   
   			//Position x (Forward)
    			IF NOT IN_xLastModalityLoadBkw AND NOT IN_xLastModalityUnloadBkw THEN
   				//Tail
   				IF TMP_dCap = 0 THEN
   					Scada_Plate[IN_iIndexArray, TMP_dCap, TMP_dLite].dTail_PosX_mm := TMP_dHeadPosition_mm - (IN_tPlate.rgtCap[TMP_dCap].dLength_cmm / 100);
   				ELSE
   					Scada_Plate[IN_iIndexArray, TMP_dCap, TMP_dLite].dTail_PosX_mm := Scada_Plate[IN_iIndexArray, TMP_dCap - 1, TMP_dLite].dTail_PosX_mm -
   					(IN_tPlate.rgtCap[TMP_dCap].dLength_cmm / 100) - (IN_tPlate.rgtCap[TMP_dCap-1].dReqGapForConv_cmm /100);	//(IN_tPlate.dGapCaps_cmm / 100);
   				END_IF;
   				//Head
   				Scada_Plate[IN_iIndexArray, TMP_dCap, TMP_dLite].dHead_PosX_mm := TMP_dHeadPosition_mm;
   				IF TMP_dCap > 0 THEN
   					Scada_Plate[IN_iIndexArray, TMP_dCap, TMP_dLite].dHead_PosX_mm := Scada_Plate[IN_iIndexArray, TMP_dCap - 1, TMP_dLite].dHead_PosX_mm -
   					(IN_tPlate.rgtCap[TMP_dCap - 1].dLength_cmm / 100) - (IN_tPlate.rgtCap[TMP_dCap-1].dReqGapForConv_cmm /100);	//(IN_tPlate.dGapCaps_cmm / 100);
   				END_IF;
   			END_IF;
   			//Position x (Backward)
   			//Head
   			IF IN_xLastModalityLoadBkw OR IN_xLastModalityUnloadBkw THEN
   				//  Head
   				IF TMP_dCap = 0 THEN
   					Scada_Plate[IN_iIndexArray, TMP_dCap, TMP_dLite].dHead_PosX_mm := TMP_dConveyorLenght - TMP_dHeadPosition_mm + (IN_tPlate.dLength_cmm / 100);
   				ELSE
   					Scada_Plate[IN_iIndexArray, TMP_dCap, TMP_dLite].dHead_PosX_mm := (TMP_dConveyorLenght - TMP_dHeadPosition_mm
   					+ (IN_tPlate.dLength_cmm / 100)) - (IN_tPlate.rgtCap[TMP_dCap - 1].dLength_cmm / 100) - (IN_tPlate.rgtCap[TMP_dCap-1].dReqGapForConv_cmm /100);	//(IN_tPlate.dGapCaps_cmm / 100);
   				END_IF;
   				//  Tail
   				IF TMP_dCap = 0 THEN
   					Scada_Plate[IN_iIndexArray, TMP_dCap, TMP_dLite].dTail_PosX_mm :=
   					Scada_Plate[IN_iIndexArray, TMP_dCap, TMP_dLite].dHead_PosX_mm - (IN_tPlate.rgtCap[TMP_dCap].dLength_cmm / 100);
   				ELSE
   					Scada_Plate[IN_iIndexArray, TMP_dCap, TMP_dLite].dTail_PosX_mm :=
   					Scada_Plate[IN_iIndexArray, TMP_dCap, TMP_dLite].dHead_PosX_mm - (IN_tPlate.rgtCap[TMP_dCap].dLength_cmm / 100);
   				END_IF;
   			END_IF;
   			//Position Y
   			//Baricentre not used, without inversion (IN Fc)
   			IF NOT IN_xYWithBaricentre AND NOT IN_xYInversionLite THEN
   				IF TMP_dLite < 1 THEN
   					Scada_Plate[IN_iIndexArray, TMP_dCap, TMP_dLite].dPositionY_mm :=
   					((TMP_dWidth_mm / 2) - (IN_tPlate.rgtCap[TMP_dCap].dWidth_cmm / 100) / 2);
   				END_IF;
   			END_IF;
   			//Baricentre not used, with inversion (IN Fc)
   			IF NOT IN_xYWithBaricentre AND IN_xYInversionLite THEN
   				IF TMP_dLite < 1 THEN
   					Scada_Plate[IN_iIndexArray, TMP_dCap, TMP_dLite].dPositionY_mm :=
   					(TMP_dWidth_mm / 2) + ((IN_tPlate.rgtCap[TMP_dCap].dWidth_cmm / 100) / 2) -
   					(IN_tPlate.rgtCap[TMP_dCap].rgtLite[TMP_dLite].dWidth_cmm / 100);
   				ELSE
   					Scada_Plate[IN_iIndexArray, TMP_dCap, TMP_dLite].dPositionY_mm := Scada_Plate[IN_iIndexArray, TMP_dCap, TMP_dLite - 1].dPositionY_mm
   					- (IN_tPlate.rgtCap[TMP_dCap].rgtLite[TMP_dLite].dWidth_cmm / 100) -
   					(IN_tPlate.rgtCap[TMP_dCap-1].dReqGapForConv_cmm /100);	//(IN_tPlate.rgtCap[TMP_dCap].dGap_cmm / 100);
   				END_IF;
   			END_IF;
   			//Baricentre used, without inversion (IN Fc)
   			IF IN_xYWithBaricentre AND NOT IN_xYInversionLite THEN
   				Scada_Plate[IN_iIndexArray, TMP_dCap, TMP_dLite].dPositionY_mm :=
   				(TMP_dWidth_mm / 2) - ((IN_tPlate.rgtCap[TMP_dCap].rgtLite[TMP_dLite].dWidth_cmm / 100) / 2)
   				+ (IN_tPlate.rgtCap[TMP_dCap].rgtLite[TMP_dLite].dBarycenter_cmm / 100);
   			END_IF;
   			//Baricentre used, with inversion (IN Fc)
   			IF IN_xYWithBaricentre AND IN_xYInversionLite THEN    //Baricentre used,  inversion
   				Scada_Plate[IN_iIndexArray, TMP_dCap, TMP_dLite].dPositionY_mm :=
   				(TMP_dWidth_mm / 2) - ((IN_tPlate.rgtCap[TMP_dCap].rgtLite[TMP_dLite].dWidth_cmm / 100) / 2)
   				- (IN_tPlate.rgtCap[TMP_dCap].rgtLite[TMP_dLite].dBarycenter_cmm / 100);
   			END_IF;
   		END_IF;
   	END_FOR;
   END_FOR;
   
END_ROUTINE
END_ADD_ON_INSTRUCTION

ADD_ON_INSTRUCTION GP_SpaceConvUtilities_V1   (* revision 1.0 *)
VAR_IN_OUT
   Conveyor : SpaceConv_Utilities; {required}
   Previus_Conveyor : SpaceConv_Utilities; {required}
   Next_Conveyor : SpaceConv_Utilities; {required}
END_VAR
VAR_INPUT
   In_dModality : DINT; {required}   // Call modality 1=GlsPos|2=PrstH|3=PrstT|4=SyncH_T|5=StartLoadForward|6=StartUnloadForward|7=PrstLoad/Unload12=PrstHInversionRun|13=PrstTInversionRun |15=StartLoadBackward|16=StartUnloadBackward
END_VAR
VAR
   TMP_dVirtualSyncroPos_cmm : DINT; {access None}
   TMP_rSP_Speed_mm_min : REAL; {access None}
   TMP_rScan_ms : REAL; {access None}
   TMP_xRunning : BOOL; {access None}
   TMP_rStepAcc_mm_min : REAL; {access None}
   TMP_rLimAcc_mm_min : REAL; {access None}
   TMP_rStepDec_mm_min : REAL; {access None}
   TMP_rLimDec_mm_min : REAL; {access None}
   TMP_dRampSpace_cmm : DINT; {access None}
   TMP_dAcc_ms2 : DINT; {access None}
   TMP_dSincrhoPhotocelPos : DINT; {access None}
   TMP_dRealSpeed : REAL; {access None}
END_VAR

ROUTINE Logic   (* structured text *)
   
   CASE In_dModality OF
       2: //Preset head position
           Conveyor.O_rHeadPosition_cmm := Conveyor.CONF_MD2_MD3_dPrstPos_cmm;
           Conveyor.O_dHeadPosition_cmm := Conveyor.CONF_MD2_MD3_dPrstPos_cmm;
   
       3: //Preset Tail position
           Conveyor.O_rTailPosition_cmm := Conveyor.CONF_MD2_MD3_dPrstPos_cmm;
           Conveyor.O_dTailPosition_cmm := Conveyor.CONF_MD2_MD3_dPrstPos_cmm;
   
       4://Glass syncrhonization
           // Calculate Ramp Space
           TMP_dAcc_ms2 := Conveyor.CONST_rAcceleration_ms2 * 1000.0;
           TMP_dRampSpace_cmm := ((Conveyor.ST_dRealSpeed_mm_min / 60) * (Conveyor.ST_dRealSpeed_mm_min / 60)) / (2 * TMP_dAcc_ms2) * 100;
           TMP_dSincrhoPhotocelPos := TMP_dRampSpace_cmm + Conveyor.CONST_dSyncroPhPosition_cmm;
           CASE Conveyor.CONST_dSyncMode OF
               0://No syncro
                   Conveyor.O_xPlateSynchronized := 1;
   
               1://Syncro on head
                   IF Conveyor.ST_OS_xSynchroPhotocellHead AND NOT (Conveyor.O_xPlateSynchronized)
                       AND Conveyor.O_dHeadPosition_cmm >= TMP_dSincrhoPhotocelPos - (Conveyor.CONST_dSyncroPhWindow_cmm / 2)
                       AND Conveyor.O_dHeadPosition_cmm <= TMP_dSincrhoPhotocelPos + (Conveyor.CONST_dSyncroPhWindow_cmm / 2) THEN
                       Conveyor.O_dHeadPosition_cmm := TMP_dSincrhoPhotocelPos;
                       Conveyor.O_rHeadPosition_cmm := Conveyor.O_dHeadPosition_cmm;
                       Conveyor.O_xPlateSynchronized := 1;
                   END_IF;
               2://Syncro on tail
                   TMP_dVirtualSyncroPos_cmm := TMP_dSincrhoPhotocelPos + Conveyor.CONF_MD4_MD6_dLength_cmm;
                   IF Conveyor.ST_OS_xSynchroPhotocellTail AND NOT (Conveyor.O_xPlateSynchronized)
                       AND Conveyor.O_dHeadPosition_cmm >= TMP_dVirtualSyncroPos_cmm - (Conveyor.CONST_dSyncroPhWindow_cmm / 2)
                       AND Conveyor.O_dHeadPosition_cmm <= TMP_dVirtualSyncroPos_cmm + (Conveyor.CONST_dSyncroPhWindow_cmm / 2) THEN
                       Conveyor.O_dHeadPosition_cmm := TMP_dVirtualSyncroPos_cmm;
                       Conveyor.O_rHeadPosition_cmm := Conveyor.O_dHeadPosition_cmm;
                       Conveyor.O_xPlateSynchronized := 1;
                   END_IF;
           END_CASE;
       5://Start load
           Conveyor.O_dHeadPosition_cmm := Previus_Conveyor.O_dHeadPosition_cmm - Previus_Conveyor.CONST_dConveyorLength_cmm;
           Conveyor.O_rHeadPosition_cmm := Conveyor.O_dHeadPosition_cmm;
           Conveyor.ST_rSpeedIncrementH_mm_min := Previus_Conveyor.ST_rSpeedIncrementH_mm_min;
           Conveyor.ST_xLastModLoadBkw := 0;
           Conveyor.ST_xLastModUnloadBkw := 0;
       6://Start unload
           Conveyor.O_dTailPosition_cmm := Conveyor.O_dHeadPosition_cmm - Conveyor.CONF_MD4_MD6_dLength_cmm;
           Conveyor.O_rTailPosition_cmm := Conveyor.O_dTailPosition_cmm;
           Conveyor.ST_xLastModLoadBkw := 0;
           Conveyor.ST_xLastModUnloadBkw := 0;
       7://Load and unload simultaneous
           TMP_dAcc_ms2 := Conveyor.CONST_rAcceleration_ms2 * 1000.0;
           TMP_dRampSpace_cmm := ((Conveyor.ST_dRealSpeed_mm_min / 60) * (Conveyor.ST_dRealSpeed_mm_min / 60)) / (2 * TMP_dAcc_ms2) * 100;
           Conveyor.O_dPresetLoadUnload_cmm := ((Conveyor.CONST_dConveyorLength_cmm + TMP_dRampSpace_cmm - Conveyor.ST_dStopLoadForseen_cmm)
           - (Previus_Conveyor.CONST_dConveyorLength_cmm - Previus_Conveyor.O_dHeadPosition_cmm)) + Conveyor.CONF_MD7_dOffset_cmm;
   
       12://Preset head position  (Inversion Run Backward Load)
           Conveyor.O_dHeadPosition_cmm := (Next_Conveyor.O_dTailPosition_cmm - Next_Conveyor.CONST_dConveyorLength_cmm) +
           Next_Conveyor.CONF_MD4_MD6_dLength_cmm;
           Conveyor.O_rHeadPosition_cmm := Conveyor.O_dHeadPosition_cmm;
           Conveyor.ST_xLastModLoadBkw := 1;
       13: //Preset Tail position (Inversion Run  Backward Unload)
          Conveyor.O_dTailPosition_cmm := Conveyor.CONST_dConveyorLength_cmm - Conveyor.O_dHeadPosition_cmm;
              Conveyor.O_rTailPosition_cmm := Conveyor.O_dTailPosition_cmm;
              Conveyor.ST_xLastModUnloadBkw := 1;
   
       15://Start Load Backward
       	IF NOT Conveyor.ST_xLastModLoadBkw THEN
           	Conveyor.O_dHeadPosition_cmm := (Next_Conveyor.O_dTailPosition_cmm-Next_Conveyor.CONST_dConveyorLength_cmm) +
           	Next_Conveyor.CONF_MD4_MD6_dLength_cmm;
           	Conveyor.O_rHeadPosition_cmm := Conveyor.O_dHeadPosition_cmm;
           	Conveyor.ST_xLastModLoadBkw := 1;
           ELSE
           	Conveyor.O_dHeadPosition_cmm := Next_Conveyor.O_dHeadPosition_cmm - Next_Conveyor.CONST_dConveyorLength_cmm;
           	Conveyor.O_rHeadPosition_cmm := Conveyor.O_dHeadPosition_cmm;
           	Conveyor.ST_rSpeedIncrementH_mm_min := Next_Conveyor.ST_rSpeedIncrementH_mm_min;
           	Conveyor.ST_xLastModLoadBkw := 1;
           END_IF;
   
       16://Start unload Backward
       	IF NOT Conveyor.ST_xLastModUnloadBkw THEN
           	Conveyor.O_dTailPosition_cmm := Conveyor.CONST_dConveyorLength_cmm - Conveyor.O_dHeadPosition_cmm;
           	Conveyor.O_rTailPosition_cmm := Conveyor.O_dTailPosition_cmm;
           	Conveyor.ST_xLastModUnloadBkw := 1;
           ELSE
           	Conveyor.O_dTailPosition_cmm := Conveyor.O_dHeadPosition_cmm - Conveyor.CONF_MD4_MD6_dLength_cmm;
           	Conveyor.O_rTailPosition_cmm := Conveyor.O_dTailPosition_cmm;
           	Conveyor.ST_xLastModUnloadBkw := 1;
   		END_IF;
   
   
   
       ELSE
           ; //Glas position
           //FEEDBACK SIMULATING TIME
           IF Conveyor.CONF_MD1_xRun OR Conveyor.CONF_MD1_xReverse THEN
               Conveyor.O_dCountFeedbackTime_ms := Conveyor.O_dCountFeedbackTime_ms - Conveyor.CONF_MD1_dScan_ms;
               IF Conveyor.O_dCountFeedbackTime_ms < 0 THEN
                   Conveyor.O_dCountFeedbackTime_ms := 0;
               END_IF;
           ELSE
               Conveyor.O_dCountFeedbackTime_ms := Conveyor.CONST_dPresetFeedbackTime_ms;
           END_IF;
   
           //Step Advancement Calculation
           //Normalize values
           Conveyor.ST_rStepAdvancementH := 0.0;
           TMP_rSP_Speed_mm_min := Conveyor.ST_dRealSpeed_mm_min;
           TMP_rScan_ms := Conveyor.CONF_MD1_dScan_ms;
           Conveyor.O_xRampInProgress := 0;
           Conveyor.O_xAccInProgress := 0;
           Conveyor.O_xDecInProgress := 0;
           TMP_xRunning := Conveyor.ST_xFeedbackRotation AND (Conveyor.CONF_MD1_xRun OR Conveyor.CONF_MD1_xReverse);
   
           //Head speed increment
           //Choose direction
           IF TMP_xRunning AND TMP_rSP_Speed_mm_min > Conveyor.ST_rSpeedIncrementH_mm_min THEN
               //Acceleration
               TMP_rStepAcc_mm_min := Conveyor.CONST_rAcceleration_ms2 * TMP_rScan_ms * 60.0;
               Conveyor.ST_rSpeedIncrementH_mm_min := Conveyor.ST_rSpeedIncrementH_mm_min + TMP_rStepAcc_mm_min;
               TMP_rLimAcc_mm_min := TMP_rSP_Speed_mm_min + TMP_rStepAcc_mm_min;
               Conveyor.O_xRampInProgress := 1;
               Conveyor.O_xAccInProgress := 1;
               IF TMP_xRunning AND Conveyor.ST_rSpeedIncrementH_mm_min > TMP_rSP_Speed_mm_min AND Conveyor.ST_rSpeedIncrementH_mm_min < TMP_rLimAcc_mm_min THEN
                   Conveyor.ST_rSpeedIncrementH_mm_min := TMP_rSP_Speed_mm_min;
               END_IF;
           ELSIF (TMP_xRunning AND TMP_rSP_Speed_mm_min < Conveyor.ST_rSpeedIncrementH_mm_min) OR (NOT (TMP_xRunning) AND Conveyor.ST_rSpeedIncrementH_mm_min > 0.0) THEN
               //Deceleration
               TMP_rStepDec_mm_min := Conveyor.CONST_rDeceleration_ms2 * TMP_rScan_ms * 60.0;
               Conveyor.ST_rSpeedIncrementH_mm_min := Conveyor.ST_rSpeedIncrementH_mm_min - TMP_rStepDec_mm_min;
               TMP_rLimDec_mm_min := TMP_rSP_Speed_mm_min - TMP_rStepDec_mm_min;
               Conveyor.O_xRampInProgress := 1;
               Conveyor.O_xDecInProgress := 1;
               IF TMP_xRunning AND Conveyor.ST_rSpeedIncrementH_mm_min < TMP_rSP_Speed_mm_min AND Conveyor.ST_rSpeedIncrementH_mm_min > TMP_rLimDec_mm_min THEN
                   Conveyor.ST_rSpeedIncrementH_mm_min := TMP_rSP_Speed_mm_min;
               END_IF;
           END_IF;
           //Erase PV_Speed if < 0
           IF Conveyor.ST_rSpeedIncrementH_mm_min < 0.0 THEN
               Conveyor.ST_rSpeedIncrementH_mm_min := 0.0;
           END_IF;
           //Tail speed increment
           //Choose direction
           IF TMP_xRunning AND TMP_rSP_Speed_mm_min > Conveyor.ST_rSpeedIncrementT_mm_min THEN
               //Acceleration
               TMP_rStepAcc_mm_min := Conveyor.CONST_rAcceleration_ms2 * TMP_rScan_ms * 60.0;
               Conveyor.ST_rSpeedIncrementT_mm_min := Conveyor.ST_rSpeedIncrementT_mm_min + TMP_rStepAcc_mm_min;
               TMP_rLimAcc_mm_min := TMP_rSP_Speed_mm_min + TMP_rStepAcc_mm_min;
               Conveyor.O_xRampInProgress := 1;
               Conveyor.O_xAccInProgress := 1;
               IF TMP_xRunning AND Conveyor.ST_rSpeedIncrementT_mm_min > TMP_rSP_Speed_mm_min AND Conveyor.ST_rSpeedIncrementT_mm_min < TMP_rLimAcc_mm_min THEN
                   Conveyor.ST_rSpeedIncrementT_mm_min := TMP_rSP_Speed_mm_min;
               END_IF;
           ELSIF (TMP_xRunning AND TMP_rSP_Speed_mm_min < Conveyor.ST_rSpeedIncrementT_mm_min) OR (NOT (TMP_xRunning) AND Conveyor.ST_rSpeedIncrementT_mm_min > 0.0) THEN
               //Deceleration
               TMP_rStepDec_mm_min := Conveyor.CONST_rDeceleration_ms2 * TMP_rScan_ms * 60.0;
               Conveyor.ST_rSpeedIncrementT_mm_min := Conveyor.ST_rSpeedIncrementT_mm_min - TMP_rStepDec_mm_min;
               TMP_rLimDec_mm_min := TMP_rSP_Speed_mm_min - TMP_rStepDec_mm_min;
               Conveyor.O_xRampInProgress := 1;
               Conveyor.O_xDecInProgress := 1;
               IF TMP_xRunning AND Conveyor.ST_rSpeedIncrementT_mm_min < TMP_rSP_Speed_mm_min AND Conveyor.ST_rSpeedIncrementT_mm_min > TMP_rLimDec_mm_min THEN
                   Conveyor.ST_rSpeedIncrementT_mm_min := TMP_rSP_Speed_mm_min;
               END_IF;
           END_IF;
           //Erase PV_Speed if < 0
           IF Conveyor.ST_rSpeedIncrementT_mm_min < 0.0 THEN
               Conveyor.ST_rSpeedIncrementT_mm_min := 0.0;
           END_IF;
           TMP_dRealSpeed := Conveyor.ST_dRealSpeed_mm_min;
           //Update Step advancement
           Conveyor.ST_rStepAdvancementH := (TMP_dRealSpeed * TMP_rScan_ms) / 600.0;
   
           //Update Step advancement
           Conveyor.ST_rStepAdvancementT := (TMP_dRealSpeed * TMP_rScan_ms) / 600.0;
   
           //POSITION CALCULATION
           //Head Position
           IF Conveyor.CONF_MD1_xHeadTracking THEN
               //Choose direction
               IF Conveyor.CONF_MD1_xReverse THEN
                   //Reverse count
                   Conveyor.O_rHeadPosition_cmm := Conveyor.O_rHeadPosition_cmm - Conveyor.ST_rStepAdvancementH;
               ELSIF Conveyor.CONF_MD1_xRun THEN
                   //Advancement
                   Conveyor.O_rHeadPosition_cmm := Conveyor.O_rHeadPosition_cmm + Conveyor.ST_rStepAdvancementH;
               END_IF;
           ELSE
               Conveyor.O_rHeadPosition_cmm := 0.0;
           END_IF;
           //Tail Position
           IF Conveyor.CONF_MD1_xTailTracking THEN
               //Choose direction
               IF Conveyor.CONF_MD1_xReverse THEN
                   //Reverse count
                   Conveyor.O_rTailPosition_cmm := Conveyor.O_rTailPosition_cmm - Conveyor.ST_rStepAdvancementT;
               ELSIF Conveyor.CONF_MD1_xRun THEN
                   //Advancement
                   Conveyor.O_rTailPosition_cmm := Conveyor.O_rTailPosition_cmm + Conveyor.ST_rStepAdvancementT;
               END_IF;
           ELSE
               Conveyor.O_rTailPosition_cmm := 0.0;
           END_IF;
           Conveyor.O_dHeadPosition_cmm := Conveyor.O_rHeadPosition_cmm;
           Conveyor.O_dTailPosition_cmm := Conveyor.O_rTailPosition_cmm;
   
   END_CASE;
   
   
   
   
   
   
END_ROUTINE
END_ADD_ON_INSTRUCTION

ADD_ON_INSTRUCTION GP_TrackingAddCap   (* revision 1.0 *)
VAR_IN_OUT
   INO_tBufferPlate : UDT_LINE_BUFFER_PLATE; {required}   // Buffer Plate
   INO_tConvoyCapToBeAdded : UDT_ConvoyCap_ZC; {required}
END_VAR
VAR_INPUT
   IN_dPosition_cmm : DINT; {access None, required}   // Cap absolute position
   IN_dRelPosition_cmm : DINT; {access None, required}   // Cap relative position
   IN_dIndConv : DINT; {access None, required}   // Index conveyor for relative position
END_VAR
VAR_OUTPUT
   OUT_xError : BOOL; {access None}   // Error
   OUT_dIndexInsertion : DINT; {access None}   // Index insertion
END_VAR
VAR_IN_OUT
   INO_tLine : UDT_LINE_TRACKING; {required}   // Tracking conveyor
END_VAR
VAR_INPUT
   IN_dEndTrackingPosition : DINT; {access None, required}   // End of tracking
END_VAR
VAR
   TMP_dCapPointer : DINT; {access None}   // Cap pointer
   TMP_dBufferSize : DINT; {access None}   // Buffer size
   TMP_dLineSize : DINT; {access None}   // Line size
END_VAR

ROUTINE Logic   (* structured text *)
   
   size(INO_tBufferPlate.rgtPlate[0],0,TMP_dBufferSize);
   size(INO_tLine.rgtTrkConv[0],0,TMP_dLineSize);
   FOR TMP_dCapPointer := 1 TO TMP_dBufferSize - 1 DO
       IF INO_tBufferPlate.rgtPlate[TMP_dCapPointer].tTracking.dLength_cmm <= 0 AND INO_tBufferPlate.rgtPlate[TMP_dCapPointer].tTracking.dPosition_cmm <= 0 THEN
   		//Copy Data To Circular Buffer
   		COP(INO_tConvoyCapToBeAdded,INO_tBufferPlate.rgtPlate[TMP_dCapPointer].tData,1);
           INO_tBufferPlate.rgtPlate[TMP_dCapPointer].tTracking.dLength_cmm := INO_tBufferPlate.rgtPlate[TMP_dCapPointer].tData.rgtCap[0].dLength_cmm;
           IF IN_dIndConv >= 0 AND IN_dIndConv < TMP_dLineSize THEN
               INO_tBufferPlate.rgtPlate[TMP_dCapPointer].tTracking.dPosition_cmm := INO_tLine.rgtTrkConv[IN_dIndConv].dStartPosition_cmm + IN_dRelPosition_cmm;
           ELSIF IN_dIndConv < 0  (*AND IN_dPosition_cmm >= dStartTrackingPosition*) AND IN_dPosition_cmm <= IN_dEndTrackingPosition THEN
               INO_tBufferPlate.rgtPlate[TMP_dCapPointer].tTracking.dPosition_cmm := IN_dPosition_cmm;   //Calculate Tracking Position
           ELSE
               OUT_xError := 1; //No conveyor D
           END_IF;
   
           EXIT;
       ELSE
           IF TMP_dCapPointer >= TMP_dBufferSize - 1 THEN
               OUT_xError := 1; //No Space in the Buffer
           END_IF;
       END_IF;
   END_FOR;// Find First Available Buffer Position
   IF NOT OUT_xError THEN
       OUT_dIndexInsertion := TMP_dCapPointer;
   ELSE
       OUT_dIndexInsertion := 0;
   END_IF;
   OUT_xError := 0;
   
END_ROUTINE
END_ADD_ON_INSTRUCTION

ADD_ON_INSTRUCTION GP_TrackingFiring   (* revision 1.0 *)
VAR_INPUT
   IN_dTarget_cmm : DINT; {access None, required}
   IN_dPosition_cmm : DINT; {access None, required}
   IN_dSpeed_mm_min : DINT; {access None, required}
   IN_dReactionTime_ms : DINT; {access None, required}
   IN_dWorkingSpace_cmm : DINT; {access None, required}
   IN_dOffsetFiringON_cmm : DINT; {access None, required}
   IN_dOffsetFiringOFF_cmm : DINT; {access None, required}
END_VAR
VAR_OUTPUT
   OUT_xPhaseON : BOOL; {access None, required}
   OUT_xFiringON : BOOL; {access None, required}
END_VAR
VAR
   TMP_dTail : DINT; {access None}
   TMP_dHead : DINT; {access None}
   TMP_dFiringOFF : DINT; {access None}
   TMP_dFiringON : DINT; {access None}
END_VAR

ROUTINE Logic   (* structured text *)
   TMP_dHead:= IN_dPosition_cmm + IN_dOffsetFiringON_cmm;
   TMP_dTail:= IN_dPosition_cmm - IN_dWorkingSpace_cmm + IN_dOffsetFiringOFF_cmm;
   TMP_dFiringON:= IN_dTarget_cmm - ((IN_dSpeed_mm_min * IN_dReactionTime_ms) / 600);
   TMP_dFiringOFF:= IN_dTarget_cmm;
   
   IF TMP_dTail >= TMP_dFiringOFF THEN
   	OUT_xFiringON := 0;
   	OUT_xPhaseON := 0;
   ELSIF TMP_dHead >= TMP_dFiringON THEN
   	OUT_xFiringON := 1;
   	OUT_xPhaseON := 1;
   ELSE
   	OUT_xFiringON := 0;
   	OUT_xPhaseON := 0;
   END_IF;
   
END_ROUTINE
END_ADD_ON_INSTRUCTION

ADD_ON_INSTRUCTION GP_TrackingFiringForConvoy   (* revision 1.0 *)
VAR_INPUT
   IN_dTarget_cmm : DINT; {access None, required}
   IN_dPosition_cmm : DINT; {access None, required}
   IN_dSpeed_mm_min : DINT; {access None, required}
   IN_dReactionTime_ms : DINT; {access None, required}
   IN_dWorkingSpace_cmm : DINT; {access None, required}
   IN_dOffsetFiringON_cmm : DINT; {access None, required}
   IN_dOffsetFiringOFF_cmm : DINT; {access None, required}
   IN_dTotalCaps : DINT; {access None, required}
END_VAR
VAR_IN_OUT
   INO_rgxActivate : DINT; {required}
   INO_rgdLengths_cmm : DINT[4]; {required}
   INO_rgdGaps_cmm : DINT[3]; {required}
END_VAR
VAR_INPUT
   IN_xContinuousMode : BOOL; {access None, required}
END_VAR
VAR_OUTPUT
   OUT_xPhaseON : BOOL; {access None, required}
   OUT_xFiringON : BOOL; {access None, required}
END_VAR
VAR
   TMP_dTail_cmm : DINT; {access None}
   TMP_dHead_cmm : DINT; {access None}
   TMP_dFiringOFF_cmm : DINT; {access None}
   TMP_dFiringON_cmm : DINT; {access None}
   TMP_dWP_cmm : DINT; {access None}
   TMP_dMinSpaceForRaise_cmm : DINT; {access None}
   TMP_rgdConvoyFiringOFF_cmm : DINT[4]; {access None}
   TMP_rgdConvoyFiringON_cmm : DINT[4]; {access None}
   TMP_dIndF : DINT; {access None}
   TMP_dDiff_cmm : DINT; {access None}
END_VAR

ROUTINE Logic   (* structured text *)
   
   IF IN_dTotalCaps < 2 THEN // not a convoy
   	TMP_dHead_cmm:= IN_dPosition_cmm + IN_dOffsetFiringON_cmm;
   	TMP_dTail_cmm:= IN_dPosition_cmm - IN_dWorkingSpace_cmm + IN_dOffsetFiringOFF_cmm;
   	TMP_dFiringON_cmm:= IN_dTarget_cmm - ((IN_dSpeed_mm_min * IN_dReactionTime_ms) / 600);
   	TMP_dFiringOFF_cmm:= IN_dTarget_cmm;
   
   	IF TMP_dTail_cmm >= TMP_dFiringOFF_cmm THEN
   		OUT_xFiringON := 0;
   		OUT_xPhaseON := 0;
   	ELSIF TMP_dHead_cmm >= TMP_dFiringON_cmm THEN
   		OUT_xFiringON := 1;
   		OUT_xPhaseON := 1;
   	ELSE
   		OUT_xFiringON := 0;
   		OUT_xPhaseON := 0;
   	END_IF;
   ELSIF ((IN_dTotalCaps > 1) AND (IN_dTotalCaps <= 4)) THEN // convoy
   	TMP_dMinSpaceForRaise_cmm := ((IN_dSpeed_mm_min * IN_dReactionTime_ms) / 600) * 2;
   	TMP_dWP_cmm := 0;
   	FOR TMP_dIndF := 0 TO IN_dTotalCaps - 1 DO
   		IF TMP_dIndF < 4 THEN
   			TMP_rgdConvoyFiringON_cmm[TMP_dIndF] := IN_dTarget_cmm - ((IN_dSpeed_mm_min * IN_dReactionTime_ms) / 600) - IN_dOffsetFiringON_cmm + TMP_dWP_cmm;
   			TMP_rgdConvoyFiringOFF_cmm[TMP_dIndF] := IN_dTarget_cmm - IN_dOffsetFiringOFF_cmm + INO_rgdLengths_cmm[TMP_dIndF] + TMP_dWP_cmm;
   			TMP_dWP_cmm := TMP_dWP_cmm + INO_rgdLengths_cmm[TMP_dIndF];
   			IF TMP_dIndF < IN_dTotalCaps - 1 THEN
   				TMP_dWP_cmm := TMP_dWP_cmm + INO_rgdGaps_cmm[TMP_dIndF];
   			END_IF;
   		END_IF;
   	END_FOR;
   	FOR TMP_dIndF := 0 TO IN_dTotalCaps - 2 DO
   		IF TMP_dIndF < 4 THEN
   			// if there is not enough space to raise the wheel before next cap anticipate raise of this cap
   			IF TMP_rgdConvoyFiringOFF_cmm[TMP_dIndF] > (TMP_rgdConvoyFiringON_cmm[TMP_dIndF + 1] - TMP_dMinSpaceForRaise_cmm) THEN
   				TMP_dDiff_cmm := TMP_rgdConvoyFiringOFF_cmm[TMP_dIndF] - TMP_rgdConvoyFiringON_cmm[TMP_dIndF + 1] + TMP_dMinSpaceForRaise_cmm;
   				TMP_rgdConvoyFiringOFF_cmm[TMP_dIndF] := (TMP_rgdConvoyFiringON_cmm[TMP_dIndF + 1] - TMP_dMinSpaceForRaise_cmm);
   				// if after anticipation there is not enough space to descend the wheel on this cap, posticipate descend on next cap
   				// and then recalculate anticipation of raise on this cap before next cap
   				IF TMP_rgdConvoyFiringOFF_cmm[TMP_dIndF] < (TMP_rgdConvoyFiringON_cmm[TMP_dIndF] + TMP_dMinSpaceForRaise_cmm) THEN
   					TMP_rgdConvoyFiringON_cmm[TMP_dIndF + 1] := TMP_rgdConvoyFiringON_cmm[TMP_dIndF + 1] + TMP_dDiff_cmm;
   					TMP_rgdConvoyFiringOFF_cmm[TMP_dIndF] := (TMP_rgdConvoyFiringON_cmm[TMP_dIndF + 1] - TMP_dMinSpaceForRaise_cmm);
   				END_IF;
   			END_IF;
   		END_IF;
   	END_FOR;
   	OUT_xFiringON := 0;
   	OUT_xPhaseON := 0;
   	INO_rgxActivate := 0;
   	IF IN_xContinuousMode THEN
   		IF TMP_rgdConvoyFiringOFF_cmm[IN_dTotalCaps - 1] >= IN_dPosition_cmm AND TMP_rgdConvoyFiringON_cmm[0] <= IN_dPosition_cmm THEN
   			OUT_xFiringON := 1;
   			OUT_xPhaseON := 1;
   		END_IF;
   	ELSE
   		IF TMP_rgdConvoyFiringOFF_cmm[IN_dTotalCaps - 1] >= IN_dPosition_cmm AND TMP_rgdConvoyFiringON_cmm[0] <= IN_dPosition_cmm THEN
   			OUT_xPhaseON := 1;
   		END_IF;
   		FOR TMP_dIndF := 0 TO IN_dTotalCaps - 1 DO
   			IF TMP_rgdConvoyFiringOFF_cmm[TMP_dIndF] >= IN_dPosition_cmm AND TMP_rgdConvoyFiringON_cmm[TMP_dIndF] <= IN_dPosition_cmm THEN
   				INO_rgxActivate.[TMP_dIndF] := 1;
   			END_IF;
   		END_FOR;
   		IF INO_rgxActivate <> 0 THEN
   			OUT_xFiringON := 1;
   		END_IF;
   	END_IF;
   END_IF;
   
END_ROUTINE
END_ADD_ON_INSTRUCTION

ADD_ON_INSTRUCTION GP_TrackingFoundDest   (* revision 1.0 *)
VAR_IN_OUT
   INO_tConvoyCap : UDT_ConvoyCap_ZC; {required}
END_VAR
VAR_INPUT
   IN_dMain : DINT; {access None, required}
   IN_dAlt : DINT; {access None, required}
   IN_d2Ch : DINT; {access None, required}
   IN_dType : DINT; {access None, required}
END_VAR
VAR_OUTPUT
   OUT_xFound : BOOL; {access None, required}
END_VAR
VAR_IN_OUT
   INO_CONST_dMaxLites : DINT; {constant, required}
END_VAR
VAR
   TMP_dLite : DINT; {access None}
   TMP_xDest : BOOL; {access None}
   TMP_dMainDestPlate : DINT; {access None}
   TMP_dAltPlate : DINT; {access None}
   TMP_d2ChPlate : DINT; {access None}
   TMP_xOnePlatePresence : BOOL; {access None}
   TMP_dMainDest : DINT; {access None}
   TMP_dAlt : DINT; {access None}
   TMP_d2Ch : DINT; {access None}
   TMP_dResult : DINT; {access None}
END_VAR

ROUTINE Logic   (* structured text *)
   
   //reset Output
   OUT_xFound := 0;
   TMP_xDest := 0;
   TMP_xOnePlatePresence := 0;
   //Mapping Variables
   TMP_dMainDest := IN_dMain;
   TMP_dAlt := IN_dAlt;
   TMP_d2Ch := IN_d2Ch;
   
   CASE IN_dType OF
       0://Search at last one Dest to IN,
               IF TMP_dMainDest >= 0 AND TMP_dMainDest <= 31 OR TMP_dAlt >= 0 AND TMP_dAlt <= 31
                   OR TMP_d2Ch >= 0 AND TMP_d2Ch <= 31 AND INO_tConvoyCap.rgtCap[0].dID <> 0 THEN
                   TMP_xDest := 0;
   
                   FOR TMP_dLite := 0 TO INO_CONST_dMaxLites - 1 DO
                       IF INO_tConvoyCap.rgtCap[0].rgtLite[TMP_dLite].dID <> 0 THEN
                           //Main
                           IF TMP_dMainDest >= 0 AND TMP_dMainDest <= 31 THEN
   							TMP_xDest := INO_tConvoyCap.rgtCap[0].rgtLite[TMP_dLite].tDestination.rgxMain.[TMP_dMainDest] OR TMP_xDest;
                           END_IF;
                           //Alt
                           IF TMP_dAlt >= 0 AND TMP_dAlt <= 31 THEN
                               TMP_xDest := INO_tConvoyCap.rgtCap[0].rgtLite[TMP_dLite].tDestination.rgxAlternative.[TMP_dAlt] OR TMP_xDest;
                           END_IF;
                           //2Chs
                           IF TMP_d2Ch >= 0 AND TMP_d2Ch <= 31 THEN
                               TMP_xDest := INO_tConvoyCap.rgtCap[0].rgtLite[TMP_dLite].tDestination.rgxSecChoice.[TMP_d2Ch] OR TMP_xDest;
                           END_IF;
                       END_IF;
                   END_FOR;
   
               END_IF;
       1://Search All Plate Dest to IN,
               IF TMP_dMainDest >= 0 AND TMP_dMainDest <= 31 OR TMP_dAlt >= 0 AND TMP_dAlt <= 31
                   OR TMP_d2Ch >= 0 AND TMP_d2Ch <= 31 AND INO_tConvoyCap.rgtCap[0].dID <> 0 THEN
                   TMP_xDest := 1;
                   FOR TMP_dLite := 0 TO INO_CONST_dMaxLites - 1 DO
                       IF INO_tConvoyCap.rgtCap[0].rgtLite[TMP_dLite].dID <> 0 THEN
                           TMP_xOnePlatePresence := 1;
                           //Main
                           IF TMP_dMainDest >= 0 AND TMP_dMainDest <= 31 THEN
                               TMP_xDest := INO_tConvoyCap.rgtCap[0].rgtLite[TMP_dLite].tDestination.rgxMain.[TMP_dMainDest] AND TMP_xDest;
                           END_IF;
                           //Alt
                           IF TMP_dAlt >= 0 AND TMP_dAlt <= 31 THEN
                               TMP_xDest := INO_tConvoyCap.rgtCap[0].rgtLite[TMP_dLite].tDestination.rgxAlternative.[TMP_dAlt] AND TMP_xDest;
                           END_IF;
                           //2Chs
                           IF TMP_d2Ch >= 0 AND TMP_d2Ch <= 31 THEN
                               TMP_xDest := INO_tConvoyCap.rgtCap[0].rgtLite[TMP_dLite].tDestination.rgxSecChoice.[TMP_d2Ch] AND TMP_xDest;
                           END_IF;
                       END_IF;
                   END_FOR;
               END_IF;
               IF NOT TMP_xOnePlatePresence THEN
                   TMP_xDest := 0;
               END_IF;
           2://Search First Plate Dest to IN,
               IF TMP_dMainDest >= 0 AND TMP_dMainDest <= 31 OR TMP_dAlt >= 0 AND TMP_dAlt <= 31
                   OR TMP_d2Ch >= 0 AND TMP_d2Ch <= 31 AND INO_tConvoyCap.rgtCap[0].dID <> 0 THEN
                   TMP_xDest := 1;
                   FOR TMP_dLite := 0 TO INO_CONST_dMaxLites - 1 DO
                       IF INO_tConvoyCap.rgtCap[0].rgtLite[TMP_dLite].dID <> 0 THEN
                           //Main
                           IF TMP_dMainDest >= 0 AND TMP_dMainDest <= 31 THEN
                               TMP_xDest := INO_tConvoyCap.rgtCap[0].rgtLite[TMP_dLite].tDestination.rgxMain.[TMP_dMainDest];
                               EXIT;
                           END_IF;
                           //Alt
                           IF TMP_dAlt >= 0 AND TMP_dAlt <= 31 THEN
                               TMP_xDest := INO_tConvoyCap.rgtCap[0].rgtLite[TMP_dLite].tDestination.rgxAlternative.[TMP_dAlt];
                               EXIT;
                           END_IF;
                           //2Chs
                           IF TMP_d2Ch >= 0 AND TMP_d2Ch <= 31 THEN
                               TMP_xDest := INO_tConvoyCap.rgtCap[0].rgtLite[TMP_dLite].tDestination.rgxSecChoice.[TMP_d2Ch];
                               EXIT;
                           END_IF;
                       END_IF;
                   END_FOR;
               END_IF;
           3://Search Last Plate Dest to IN,
               IF TMP_dMainDest >= 0 AND TMP_dMainDest <= 31 OR TMP_dAlt >= 0 AND TMP_dAlt <= 31
                   OR TMP_d2Ch >= 0 AND TMP_d2Ch <= 31 AND INO_tConvoyCap.rgtCap[0].dID <> 0 THEN
                   TMP_xDest := 1;
                   FOR TMP_dLite := INO_CONST_dMaxLites - 1 TO 0  BY -1 DO
                       IF INO_tConvoyCap.rgtCap[0].rgtLite[TMP_dLite].dID <> 0 THEN
                           //Main
                           IF TMP_dMainDest >= 0 AND TMP_dMainDest <= 31 THEN
                               TMP_xDest := INO_tConvoyCap.rgtCap[0].rgtLite[TMP_dLite].tDestination.rgxMain.[TMP_dMainDest];
                               EXIT;
                           END_IF;
                           //Alt
                           IF TMP_dAlt >= 0 AND TMP_dAlt <= 31 THEN
                               TMP_xDest := INO_tConvoyCap.rgtCap[0].rgtLite[TMP_dLite].tDestination.rgxAlternative.[TMP_dAlt];
                               EXIT;
                           END_IF;
                           //2Chs
                           IF TMP_d2Ch >= 0 AND TMP_d2Ch <= 31 THEN
                               TMP_xDest := INO_tConvoyCap.rgtCap[0].rgtLite[TMP_dLite].tDestination.rgxSecChoice.[TMP_d2Ch];
                               EXIT;
                           END_IF;
                       END_IF;
                   END_FOR;
               END_IF;
           10://Search at last one Dest to IN mask Version
               TMP_xDest := 0;
               FOR TMP_dLite := 0 TO INO_CONST_dMaxLites - 1 DO
                   //Main
                   IF TMP_dMainDest >= 0 THEN
                       TMP_dMainDestPlate := INO_tConvoyCap.rgtCap[0].rgtLite[TMP_dLite].tDestination.rgxMain;
                       TMP_dResult := TMP_dMainDestPlate AND TMP_dMainDestPlate;
                       TMP_xDest := TMP_dResult <> 0 OR TMP_xDest;
                   END_IF;
                   //Alt
                   IF TMP_dAlt >= 0 THEN
                       TMP_dAltPlate := INO_tConvoyCap.rgtCap[0].rgtLite[TMP_dLite].tDestination.rgxAlternative;
                       TMP_dResult := TMP_dAltPlate AND TMP_dAlt;
                       TMP_xDest := TMP_dResult <> 0 OR TMP_xDest;
                   END_IF;
                   //SecondChoise
                   IF TMP_d2Ch >= 0 THEN
                       TMP_d2ChPlate := INO_tConvoyCap.rgtCap[0].rgtLite[TMP_dLite].tDestination.rgxSecChoice;
                       TMP_dResult := TMP_d2ChPlate AND TMP_d2Ch;
                       TMP_xDest := TMP_dResult <> 0 OR TMP_xDest;
                   END_IF;
               END_FOR;
   
         11:// 11:Search All Plate Dest to IN mask Version
               TMP_xDest := 1;
               FOR TMP_dLite := 0 TO INO_CONST_dMaxLites - 1 DO
                   IF INO_tConvoyCap.rgtCap[0].rgtLite[TMP_dLite].dID <> 0 THEN
                       TMP_xOnePlatePresence := 1;
                       //Main
                       IF TMP_dMainDest >= 0 THEN
                           TMP_dMainDestPlate := INO_tConvoyCap.rgtCap[0].rgtLite[TMP_dLite].tDestination.rgxMain;
                           TMP_dResult := TMP_dMainDestPlate AND TMP_dMainDestPlate;
                           TMP_xDest := TMP_dResult <> 0 AND TMP_xDest;
                       END_IF;
                       //Alt
                       IF TMP_dAlt >= 0 THEN
                           TMP_dAltPlate := INO_tConvoyCap.rgtCap[0].rgtLite[TMP_dLite].tDestination.rgxAlternative;
                           TMP_dResult := TMP_dAltPlate AND TMP_dAlt;
                           TMP_xDest := TMP_dResult <> 0 AND TMP_xDest;
                       END_IF;
                       //SecondChoise
                       IF TMP_d2Ch >= 0 THEN
                        	TMP_d2ChPlate := INO_tConvoyCap.rgtCap[0].rgtLite[TMP_dLite].tDestination.rgxSecChoice;
                           TMP_dResult := TMP_d2ChPlate AND TMP_d2Ch;
                           TMP_xDest := TMP_dResult <> 0 AND TMP_xDest;
                       END_IF;
                   END_IF;
               END_FOR;
               IF NOT TMP_xOnePlatePresence THEN
                   TMP_xDest := 0;
               END_IF;
           12: // 12:Search first lite to IN
               TMP_xDest := 0;
               FOR TMP_dLite := 0 TO INO_CONST_dMaxLites - 1 DO
                   IF INO_tConvoyCap.rgtCap[0].rgtLite[TMP_dLite].dID <> 0 THEN
                       //Main
                       IF TMP_dMainDest >= 0 THEN
                           TMP_dMainDestPlate := INO_tConvoyCap.rgtCap[0].rgtLite[TMP_dLite].tDestination.rgxMain;
                           TMP_dResult := TMP_dMainDestPlate AND TMP_dMainDestPlate;
                           TMP_xDest := TMP_dResult <> 0;
                           EXIT;
                       END_IF;
                       //Alt
                       IF TMP_dAlt >= 0 THEN
                           TMP_dAltPlate := INO_tConvoyCap.rgtCap[0].rgtLite[TMP_dLite].tDestination.rgxAlternative;
                           TMP_dResult := TMP_dAltPlate AND TMP_dAlt;
                           TMP_xDest := TMP_dResult <> 0;
                           EXIT;
                       END_IF;
                       //SecondChoise
                       IF TMP_d2Ch >= 0 THEN
                           TMP_d2ChPlate := INO_tConvoyCap.rgtCap[0].rgtLite[TMP_dLite].tDestination.rgxSecChoice;
                           TMP_dResult := TMP_d2ChPlate AND TMP_d2Ch;
                           TMP_xDest := TMP_dResult <> 0;
                           EXIT;
                       END_IF;
                   END_IF;
               END_FOR;
           13: // 13:Search last lite to IN
               FOR TMP_dLite := INO_CONST_dMaxLites - 1 TO 0  BY -1 DO
                   IF INO_tConvoyCap.rgtCap[0].rgtLite[TMP_dLite].dID <> 0  THEN
                       IF TMP_dMainDest >= 0 THEN
                           TMP_dMainDestPlate := INO_tConvoyCap.rgtCap[0].rgtLite[TMP_dLite].tDestination.rgxMain;
                           TMP_dResult := TMP_dMainDestPlate AND TMP_dMainDestPlate;
                           TMP_xDest := TMP_dResult <> 0 ;
                           EXIT;
                           //Alt
                           IF TMP_dAlt >= 0 THEN
                               TMP_dAltPlate := INO_tConvoyCap.rgtCap[0].rgtLite[TMP_dLite].tDestination.rgxAlternative;
                               TMP_dResult := TMP_dAltPlate AND TMP_dAlt;
                               TMP_xDest := TMP_dResult <> 0;
                               EXIT;
                           END_IF;
                           //SecondChoise
                           IF TMP_d2Ch >= 0 THEN
                               TMP_d2ChPlate := INO_tConvoyCap.rgtCap[0].rgtLite[TMP_dLite].tDestination.rgxSecChoice;
                               TMP_dResult := TMP_d2ChPlate AND TMP_d2Ch;
                               TMP_xDest := TMP_dResult <> 0;
                               EXIT;
                           END_IF;
                       END_IF;
                   END_IF;
               END_FOR;
   
           ELSE  // Statement section ELSE
               ;
    END_CASE;
   
   OUT_xFound := TMP_xDest;
END_ROUTINE
END_ADD_ON_INSTRUCTION

ADD_ON_INSTRUCTION GP_TrackingGetFirstPlateInConveyor   (* revision 1.0 *)
VAR_IN_OUT
   INO_tTrkConv : UDT_ConveyorTracking; {required}   // Tracking conveyor
END_VAR
VAR_INPUT
   IN_NumCapsConveyor : DINT; {access Read Only, required}   // Max num caps for conveyor
END_VAR
VAR_OUTPUT
   OUT_dIndex : DINT; {access Read Only, required}   // Plate Index
   OUT_dHeadPos : DINT; {access Read Only, required}   // Head position of first plate in conveyor
END_VAR
VAR
   TMP_dIndCap : DINT; {access None}
END_VAR

ROUTINE Logic   (* structured text *)
   
   OUT_dIndex := 0;
   OUT_dHeadPos := 0;
   
   //Search The index of Cap
   FOR TMP_dIndCap := 0 TO IN_NumCapsConveyor - 1 DO
       //Search cap max head position
       IF INO_tTrkConv.Cap[TMP_dIndCap].dHeadPos_cmm > OUT_dHeadPos THEN
           OUT_dHeadPos := INO_tTrkConv.Cap[TMP_dIndCap].dHeadPos_cmm;
   		OUT_dIndex := INO_tTrkConv.Cap[TMP_dIndCap].dPointer;
       END_IF;
   END_FOR;
   
END_ROUTINE
END_ADD_ON_INSTRUCTION
